// TIA Portal project "management parcare auto" (V17) (continued)
      ProcessValue <- "Status2"
   IOField "I/O field_77" at 1105,395 size 126x54; FormatPattern 9
      ProcessValue <- "Status3"
   IOField "I/O field_78" at 1105,445 size 126x54; FormatPattern 9
      ProcessValue <- "Status4"
   IOField "I/O field_79" at 1105,495 size 126x54; FormatPattern 9
      ProcessValue <- "Status5"
   IOField "I/O field_80" at 1105,545 size 126x54; FormatPattern 9
      ProcessValue <- "Status6"
   IOField "I/O field_81" at 1105,595 size 126x54; FormatPattern 9
      ProcessValue <- "Status7"
   IOField "I/O field_82" at 1105,645 size 126x54; FormatPattern 9
      ProcessValue <- "Status8"
   IOField "I/O field_83" at 1105,695 size 126x54; FormatPattern 9
      ProcessValue <- "Status9"
   IOField "I/O field_84" at 1105,745 size 126x54; FormatPattern 9
      ProcessValue <- "Status10"
   IOField "I/O field_85" at 1227,345 size 177x54; FormatPattern 9999999999999999999999999999999999999999
      ProcessValue <- "EntryTime2"
   IOField "I/O field_86" at 1227,395 size 177x54; FormatPattern 9999999999999999999999999999999999999999
      ProcessValue <- "EntryTime3"
   IOField "I/O field_87" at 1227,445 size 177x54; FormatPattern 9999999999999999999999999999999999999999
      ProcessValue <- "EntryTime4"
   IOField "I/O field_88" at 1227,495 size 177x54; FormatPattern 9999999999999999999999999999999999999999
      ProcessValue <- "EntryTime5"
   IOField "I/O field_89" at 1227,545 size 177x54; FormatPattern 9999999999999999999999999999999999999999
      ProcessValue <- "EntryTime6"
   IOField "I/O field_90" at 1227,595 size 177x54; FormatPattern 9999999999999999999999999999999999999999
      ProcessValue <- "EntryTime7"
   IOField "I/O field_91" at 1227,645 size 177x54; FormatPattern 9999999999999999999999999999999999999999
      ProcessValue <- "EntryTime8"
   IOField "I/O field_92" at 1227,695 size 177x54; FormatPattern 9999999999999999999999999999999999999999
      ProcessValue <- "EntryTime9"
   IOField "I/O field_93" at 1227,745 size 177x54; FormatPattern 9999999999999999999999999999999999999999
      ProcessValue <- "EntryTime10"
   IOField "I/O field_94" at 1400,344 size 165x54; FormatPattern 9999999999999999999999999999999999999999
      ProcessValue <- "EntryDate2"
   IOField "I/O field_95" at 1401,394 size 165x54; FormatPattern 9999999999999999999999999999999999999999
      ProcessValue <- "EntryDate3"
   IOField "I/O field_96" at 1401,444 size 165x54; FormatPattern 9999999999999999999999999999999999999999
      ProcessValue <- "EntryDate4"
   IOField "I/O field_97" at 1401,494 size 165x54; FormatPattern 9999999999999999999999999999999999999999
      ProcessValue <- "EntryDate5"
   IOField "I/O field_98" at 1401,545 size 165x54; FormatPattern 9999999999999999999999999999999999999999
      ProcessValue <- "EntryDate6"
   IOField "I/O field_99" at 1401,595 size 165x54; FormatPattern 9999999999999999999999999999999999999999
      ProcessValue <- "EntryDate7"
   IOField "I/O field_100" at 1401,645 size 165x54; FormatPattern 9999999999999999999999999999999999999999
      ProcessValue <- "EntryDate8"
   IOField "I/O field_101" at 1401,695 size 165x54; FormatPattern 9999999999999999999999999999999999999999
      ProcessValue <- "EntryDate9"
   IOField "I/O field_102" at 1401,745 size 165x54; FormatPattern 9999999999999999999999999999999999999999
      ProcessValue <- "EntryDate10"
   IOField "I/O field_103" at 1562,344 size 164x54; FormatPattern 9999999999999999999999999999999999999999
      ProcessValue <- "ExitTime2"
   IOField "I/O field_104" at 1562,394 size 164x54; FormatPattern 9999999999999999999999999999999999999999
      ProcessValue <- "ExitTime3"
   IOField "I/O field_105" at 1562,444 size 164x54; FormatPattern 9999999999999999999999999999999999999999
      ProcessValue <- "ExitTime4"
   IOField "I/O field_106" at 1562,494 size 164x54; FormatPattern 9999999999999999999999999999999999999999
      ProcessValue <- "ExitTime5"
   IOField "I/O field_107" at 1562,545 size 164x54; FormatPattern 9999999999999999999999999999999999999999
      ProcessValue <- "ExitTime6"
   IOField "I/O field_108" at 1562,595 size 164x54; FormatPattern 9999999999999999999999999999999999999999
      ProcessValue <- "ExitTime7"
   IOField "I/O field_109" at 1562,645 size 164x54; FormatPattern 9999999999999999999999999999999999999999
      ProcessValue <- "ExitTime8"
   IOField "I/O field_110" at 1562,695 size 164x54; FormatPattern 9999999999999999999999999999999999999999
      ProcessValue <- "ExitTime9"
   IOField "I/O field_111" at 1562,745 size 164x54; FormatPattern 9999999999999999999999999999999999999999
      ProcessValue <- "ExitTime10"
   IOField "I/O field_112" at 1723,344 size 163x54; FormatPattern 9999999999999999999999999999999999999999
      ProcessValue <- "ExitDate2"
   IOField "I/O field_113" at 1723,394 size 163x54; FormatPattern 9999999999999999999999999999999999999999
      ProcessValue <- "ExitDate3"
   IOField "I/O field_114" at 1723,444 size 163x54; FormatPattern 9999999999999999999999999999999999999999
      ProcessValue <- "ExitDate4"
   IOField "I/O field_115" at 1723,494 size 163x54; FormatPattern 9999999999999999999999999999999999999999
      ProcessValue <- "ExitDate5"
   IOField "I/O field_116" at 1723,544 size 163x54; FormatPattern 9999999999999999999999999999999999999999
      ProcessValue <- "ExitDate6"
   IOField "I/O field_117" at 1723,594 size 163x54; FormatPattern 9999999999999999999999999999999999999999
      ProcessValue <- "ExitDate7"
   IOField "I/O field_118" at 1723,644 size 163x54; FormatPattern 9999999999999999999999999999999999999999
      ProcessValue <- "ExitDate8"
   IOField "I/O field_119" at 1723,694 size 163x54; FormatPattern 9999999999999999999999999999999999999999
      ProcessValue <- "ExitDate9"
   IOField "I/O field_120" at 1723,744 size 163x54; FormatPattern 9999999999999999999999999999999999999999
      ProcessValue <- "ExitDate10"
   TextField "Text field_4" at 994,221 size 165x119; Text 'Car number'
   TextField "Text field_6" at 11,130 size 645x121; Text 'Temporar data'
   TextField "Text field_8" at 978,132 size 901x121; Text 'Permanent data'

screen "Statistics" 1920x1080
   on GenerateScreen: "Statistica_masini_total"()
   Button "Button_3" at 608,973 size 194x96; TextOff 'Statistics'
      on Press: ActivateScreen("Statistics", 0)
   Button "Button_8" at 408,973 size 194x96; TextOff 'Parking history'
      on Press: ActivateScreen("Parking history", 0)
   Button "Button_1" at 208,973 size 194x96; TextOff 'Alarms'
      on Press: ActivateScreen("Alarms", 0)
   Button "Button_2" at 9,972 size 194x96; TextOff 'Home / Ecran principal'
      on Press: ActivateScreen("Home", 0)
   GraphicView "Graphic view_2" at 28,12 size 394x64; Picture "Siemens_AG_logo.svg"
   Button "Button_4" at 1748,4 size 170x79; TextOff 'Exit / Iesire'
      on Press: StopRuntime(0)
   TextField "Text field_1" at 184,382 size 485x109; Text 'Number of cars:'
   TextField "Text field_2" at 794,230 size 49x81; Text 'Text'
   TextField "Text field_3" at 615,147 size 581x176; Text 'STATISTICS'
   TextField "Text field_4" at 164,210 size 1445x179; Text 'Choose a date(yy-mm-dd) to find out the number of cars on that day:'
   TextField "Text field_5" at 166,452 size 1589x179; Text 'Choose an interval to find out the number of cars in that period of time:'
   IOField "I/O field_1" at 316,328 size 178x62; FormatPattern ??????????
      on OnFinishInput: "Statistica_masini_zi"()
      ProcessValue <- "filtrare_dupa_data"
   IOField "I/O field_2" at 641,404 size 128x68; FormatPattern 99999
      ProcessValue <- "Numar_masini_ziuaX"
   TextField "Text field_6" at 512,561 size 26x62; Text '-'
   IOField "I/O field_4" at 312,569 size 188x62; FormatPattern ??????????
      ProcessValue <- "Interval1_date"
   IOField "I/O field_3" at 566,568 size 188x62; FormatPattern ??????????
      on OnFinishInput: "Statistica_masini_pe_interval"()
      ProcessValue <- "Interval2_date"
   TextField "Text field_7" at 166,621 size 485x109; Text 'Number of cars:'
   IOField "I/O field_5" at 615,647 size 128x68; FormatPattern 99999
      ProcessValue <- "nr_masini_interval"
   TextField "Text field_8" at 262,783 size 725x133; Text 'Total number of cars:'
   IOField "I/O field_6" at 1006,829 size 204x52; FormatPattern 9999999
      ProcessValue <- "nr_total_masini"

VB script "Insert_to_database"
   'RdyToLog= un tagg care se face 1 atunci cand butonul entry de pe HMI(nu runtime) este activat, devine trigger pentru a rula scriptul
   SmartTags("Verficare_rulareScriptInsr")=0
   If (SmartTags("RdyToLog")=True) And (SmartTags("04_DB_MarkersAuto_car status_1")=True Or SmartTags("04_DB_MarkersAuto_car status_2")=True Or SmartTags("04_DB_MarkersAuto_car status_3")=True Or SmartTags("04_DB_MarkersAuto_car status_4")=True Or SmartTags("04_DB_MarkersAuto_car status_5")=True Or SmartTags("04_DB_MarkersAuto_car status_6")=True Or SmartTags("04_DB_MarkersAuto_car status_7")=True Or SmartTags("04_DB_MarkersAuto_car status_8")=True Or SmartTags("04_DB_MarkersAuto_car status_9")=True Or SmartTags("04_DB_MarkersAuto_car status_10")=True ) Then
   
   Dim rs,con
   Dim nrMasina, statusMasina, oraIntrare,dataIntrare,oraIesire,dataIesire,dsValueEntry,dsValueExit
   
   
   'se ia nr de masina introdus de utilizator
   Set nrMasina= SmartTags("02_DB_HMI_Buttons_nr_masina")
   
   'se seteaza statusul masinii in functie de ce loc a ocupat
   If SmartTags("04_DB_MarkersAuto_car status_1")=True Then
   	statusMasina= 1
   End If
   
   If SmartTags("04_DB_MarkersAuto_car status_2")=True  Then
   	statusMasina=1
   End If
   
   If SmartTags("04_DB_MarkersAuto_car status_3")=True Then
   	statusMasina=1
   End If
   
   If SmartTags("04_DB_MarkersAuto_car status_4")=True Then
   	statusMasina=1
   End If
   
   If SmartTags("04_DB_MarkersAuto_car status_5")=True Then
   	statusMasina=1
   End If
   
   If SmartTags("04_DB_MarkersAuto_car status_6")=True Then
   	statusMasina=1
   End If
   
   If SmartTags("04_DB_MarkersAuto_car status_7")=True Then
   	statusMasina=1
   End If
   
   If SmartTags("04_DB_MarkersAuto_car status_8")=True Then
   	statusMasina=1
   End If
   
   If SmartTags("04_DB_MarkersAuto_car status_9")=True Then
   	statusMasina=1
   End If
   
   If  SmartTags("04_DB_MarkersAuto_car status_10")=True Then
   	statusMasina=1
   End If
   
   
   
   'Dim Timp
   'Timp = Time
   'Dim TimpStamp
   Dim dtsnow
   Dim dd, mm, yy, hh, nn, ss
   Dim DataValue, TimpValue
   
   'atunci cand se intra in parcare, se ia ora si data intrarii
   If SmartTags("11_DB_Inputs_i0.0")=True Then
   ' Obține data și ora curentă
   dtsnow = Now()
   dd = Right("00" & Day(dtsnow), 2)
   mm = Right("00" & Month(dtsnow), 2)
   yy = Year(dtsnow)
   
   hh = Right("00" & Hour(dtsnow), 2)
   nn = Right("00" & Minute(dtsnow), 2)
   ss = Right("00" & Second(dtsnow), 2)
   
   'Build the date string in the format yyyy-mm-dd
   dataIntrare = yy & "-" & mm & "-" & dd
   'Build the time string in the format hh:mm:ss
   oraIntrare = hh & ":" & nn & ":" & ss
   dsValueEntry=dataIntrare &" "& oraIntrare
   End If
   
   'atunci cand se plateste se ia ora si data iesirii
   If SmartTags("02_DB_HMI_Buttons_pay")=True Then
   ' Obține data și ora curentă
   dtsnow = Now()
   dd = Right("00" & Day(dtsnow), 2)
   mm = Right("00" & Month(dtsnow), 2)
   yy = Year(dtsnow)
   
   hh = Right("00" & Hour(dtsnow), 2)
   nn = Right("00" & Minute(dtsnow), 2)
   ss = Right("00" & Second(dtsnow), 2)
   
   'Build the date string in the format dd-mm-yyyy
   dataIesire = yy & "-" & mm & "-" & dd
   'Build the time string in the format hh:mm:ss
   oraIesire = hh & ":" & nn & ":" & ss
   dsValueExit=dataIesire & " " &oraIesire
   
   End If
   
   'conexiune baza de date si inserare
   Set con=CreateObject("adodb.connection")
   Set rs=CreateObject("adodb.recordset")
   
   con.open"Driver={MySQL ODBC 8.0 Unicode Driver};Server=localhost:3306;Database=parkingcar;User=root;Password=;Option=3;"
   Dim rezultate,rez
   rez="INSERT INTO parkingcar.permanent(NrInm,StatusMasina,OraIntrare,DataIntrare,OraIesire,DataIesire,DataOraEntry,DataOraExit) VALUES ('" & nrMasina & "', '" & statusMasina & "', '" & oraIntrare & "','" & dataIntrare & "','" & oraIesire & "','" & dataIesire & "', '" & dsValueEntry &"','"& dsValueExit &"')"
   rezultate= "INSERT INTO parkingcar.temporar(NrInm,StatusMasina,OraIntrare,DataIntrare,OraIesire,DataIesire,DataOraIntr,DataOraIesire) VALUES ('" & nrMasina & "', '" & statusMasina & "', '" & oraIntrare & "','" & dataIntrare & "','" & oraIesire & "','" & dataIesire & "', '" & dsValueEntry &"','"& dsValueExit &"')"
   rs.open rezultate,con
   rs.open rez,con
   con.Close
   End If
   
   SmartTags("Verficare_rulareScriptInsr")=1

VB script "EditDataRecord"
   'Tip:
   ' 1. Use the <CTRL+SPACE> or <CTRL+I> shortcut to open a list of all objects and functions
   ' 2. Write the code using the HMI Runtime object.
   '  Example: HmiRuntime.Screens("Screen_1").
   ' 3. Use the <CTRL+J> shortcut to create an object reference.
   'Write the code as of this position:
   
   
   If SmartTags("RdyToUpdate")=True Then
   Dim nrMasina,statusMasina, oraIesire,dataIesire
   Dim con,rs
   
   'se ia nr de masina folosit pentru a iesi din parcare
   Set nrMasina=SmartTags("02_DB_HMI_Buttons_nrMasina_iesire")
   
   If SmartTags("04_DB_MarkersAuto_car status_1")=False Then
   	statusMasina= 0
   End If
   
   If SmartTags("04_DB_MarkersAuto_car status_2")=False  Then
   	statusMasina=0
   End If
   
   If SmartTags("04_DB_MarkersAuto_car status_3")=False Then
   	statusMasina=0
   End If
   
   If SmartTags("04_DB_MarkersAuto_car status_4")=False Then
   	statusMasina=0
   End If
   
   If SmartTags("04_DB_MarkersAuto_car status_5")=False Then
   	statusMasina=0
   End If
   
   If SmartTags("04_DB_MarkersAuto_car status_6")=False Then
   	statusMasina=0
   End If
   
   If SmartTags("04_DB_MarkersAuto_car status_7")=False Then
   	statusMasina=0
   End If
   
   If SmartTags("04_DB_MarkersAuto_car status_8")=False Then
   	statusMasina=0
   End If
   
   If SmartTags("04_DB_MarkersAuto_car status_9")=False Then
   	statusMasina=0
   End If
   
   If  SmartTags("04_DB_MarkersAuto_car status_10")=False Then
   	statusMasina=0
   End If
   
   
   Dim dtsnow
   Dim dd, mm, yy, hh, nn, ss
   Dim DataValue, TimpValue,dsValueExit
   
   'atunci cand se plateste se ia ora si data iesirii
   If SmartTags("11_DB_Inputs_i1.0")=True Then
   ' Obține data și ora curentă
   dtsnow = Now()
   dd = Right("00" & Day(dtsnow), 2)
   mm = Right("00" & Month(dtsnow), 2)
   yy = Year(dtsnow)
   
   hh = Right("00" & Hour(dtsnow), 2)
   nn = Right("00" & Minute(dtsnow), 2)
   ss = Right("00" & Second(dtsnow), 2)
   
   'Build the date string in the format dd-mm-yyyy
   dataIesire = yy & "-" & mm & "-" & dd
   'Build the time string in the format hh:mm:ss
   oraIesire = hh & ":" & nn & ":" & ss
   dsValueExit=dataIesire &" " &oraIesire
   End If
   
   'conxiune baza de date si editare ora iesire si statusul
   Set con=CreateObject("adodb.connection")
   Set rs=CreateObject("adodb.recordset")
   
   con.open"Driver={MySQL ODBC 8.0 Unicode Driver};Server=localhost:3306;Database=parkingcar;User=root;Password=;Option=3;"
   Dim rezultate,rez
   rez="UPDATE parkingcar.permanent SET StatusMasina='" & statusMasina &"',OraIesire='" & oraIesire & "',DataIesire='" & dataIesire &"',DataOraExit='"& dsValueExit &"' WHERE NrInm='" & nrMasina &"' "
   rezultate= "UPDATE parkingcar.temporar SET StatusMasina='" & statusMasina &"',OraIesire='" & oraIesire & "',DataIesire='" & dataIesire &"', DataOraIesire='"& dsValueExit &"' WHERE NrInm='" & nrMasina &"' "
   rs.open rezultate,con
   rs.open rez,con
   con.Close
   
   End If

VB script "Delete_from_database"
   'Tip:
   ' 1. Use the <CTRL+SPACE> or <CTRL+I> shortcut to open a list of all objects and functions
   ' 2. Write the code using the HMI Runtime object.
   '  Example: HmiRuntime.Screens("Screen_1").
   ' 3. Use the <CTRL+J> shortcut to create an object reference.
   'Write the code as of this position:
   
   If SmartTags("RdyToDelete")=True Then
   	
   Dim con,rs
   
   Set con=CreateObject("adodb.connection")
   Set rs=CreateObject("adodb.recordset")
   
   con.open"Driver={MySQL ODBC 8.0 Unicode Driver};Server=localhost:3306;Database=parkingcar;User=root;Password=;Option=3;"
   Dim rezultate
   rezultate= "DELETE FROM parkingcar.temporar WHERE StatusMasina= '0'"
   rs.open rezultate,con
   con.Close
   End If

VB script "Statistica_masini_zi"
   'Tip:
   ' 1. Use the <CTRL+SPACE> or <CTRL+I> shortcut to open a list of all objects and functions
   ' 2. Write the code using the HMI Runtime object.
   '  Example: HmiRuntime.Screens("Screen_1").
   ' 3. Use the <CTRL+J> shortcut to create an object reference.
   'Write the code as of this position:
   
   Dim con,rs 
   Set con=CreateObject("ADODB.Connection")
   Set rs= CreateObject("adodb.recordset")
   
   con.Open "DRIVER={MySQL ODBC 8.0 Unicode Driver};Server=localhost:3306;Database=parkingcar;User=root;Password=;Option=3;"
   rs.open "SELECT  COUNT(* ) AS NumarMasini FROM permanent WHERE DataIntrare = '" & SmartTags("filtrare_dupa_data")&"' ",con
   SmartTags("Numar_masini_ziuaX")=rs.Fields(0)
   Set con=Nothing

VB script "Statistica_masini_pe_interval"
   'Tip:
   ' 1. Use the <CTRL+SPACE> or <CTRL+I> shortcut to open a list of all objects and functions
   ' 2. Write the code using the HMI Runtime object.
   '  Example: HmiRuntime.Screens("Screen_1").
   ' 3. Use the <CTRL+J> shortcut to create an object reference.
   'Write the code as of this position:
   Dim con,rs 
   Set con=CreateObject("ADODB.Connection")
   Set rs= CreateObject("adodb.recordset")
   
   con.Open "DRIVER={MySQL ODBC 8.0 Unicode Driver};Server=localhost:3306;Database=parkingcar;User=root;Password=;Option=3;"
   rs.open "SELECT  COUNT(* ) AS NumarMasini FROM permanent WHERE DataIntrare >= '" & SmartTags("Interval1_date") &"' AND DataIntrare <= '" & SmartTags("Interval2_date") &"' ",con
   SmartTags("nr_masini_interval")=rs.Fields(0)

VB script "Statistica_masini_total"
   'Tip:
   ' 1. Use the <CTRL+SPACE> or <CTRL+I> shortcut to open a list of all objects and functions
   ' 2. Write the code using the HMI Runtime object.
   '  Example: HmiRuntime.Screens("Screen_1").
   ' 3. Use the <CTRL+J> shortcut to create an object reference.
   'Write the code as of this position:
   
   Dim con,rs 
   Set con=CreateObject("ADODB.Connection")
   Set rs= CreateObject("adodb.recordset")
   
   con.Open "DRIVER={MySQL ODBC 8.0 Unicode Driver};Server=localhost:3306;Database=parkingcar;User=root;Password=;Option=3;"
   rs.open "SELECT  COUNT(* ) AS NumarMasini FROM permanent",con
   SmartTags("nr_total_masini")=rs.Fields(0)

VB script "Read_fromTEMP"
   'Tip:
   ' 1. Use the <CTRL+SPACE> or <CTRL+I> shortcut to open a list of all objects and functions
   ' 2. Write the code using the HMI Runtime object.
   '  Example: HmiRuntime.Screens("Screen_1").
   ' 3. Use the <CTRL+J> shortcut to create an object reference.
   'Write the code as of this position:
   Dim con,rs
   ' Creează obiectul pentru conexiunea la bază de date
   Set con = CreateObject("ADODB.Connection")
   Set rs=CreateObject("adodb.recordset")
    
   ' Deschide conexiunea la bază de date
   con.Open "DRIVER={MySQL ODBC 8.0 Unicode Driver};Server=localhost:3306;Database=parkingcar;User=root;Password=;Option=3;"
   rs.open "SELECT * FROM temporar ORDER BY NrInm ASC ",con
   rs.MoveFirst
   Dim i
   i=1
   While Not rs.EOF
   SmartTags("NrMasina"& i)=rs.Fields("NrInm")
   SmartTags("CarStatus"& i)=rs.Fields("StatusMasina")
   SmartTags("OraIntrare"& i)=rs.Fields("DataOraIntr")
   SmartTags("DataIntrare"& i)=rs.Fields("DataOraIntr")
   rs.MoveNext
   i=i+1
   Wend
   
   If rs.EOF Then
   	rs.Close
   	con.Close
   End If

VB script "Read_fromPerm"
   'Tip:
   ' 1. Use the <CTRL+SPACE> or <CTRL+I> shortcut to open a list of all objects and functions
   ' 2. Write the code using the HMI Runtime object.
   '  Example: HmiRuntime.Screens("Screen_1").
   ' 3. Use the <CTRL+J> shortcut to create an object reference.
   'Write the code as of this position:
   
   Dim con,rs
   ' Creează obiectul pentru conexiunea la bază de date
   Set con = CreateObject("ADODB.Connection")
   Set rs=CreateObject("adodb.recordset")
    Dim exittime
    exittime="00-00-00 00:00:00"
   ' Deschide conexiunea la bază de date
   con.Open "DRIVER={MySQL ODBC 8.0 Unicode Driver};Server=localhost:3306;Database=parkingcar;User=root;Password=;Option=3;"
   rs.open "SELECT * FROM permanent ORDER BY DataIntrare DESC",con
   rs.MoveFirst
   Dim i
   'Please replace all sequences which are enclosed with '_' by your own code.
   For  i= 1 To 10
   SmartTags("CarNumber"& i)=rs.Fields("NrInm")
   SmartTags("Status"& i)=rs.Fields("StatusMasina")
   SmartTags("EntryTime"& i)=rs.Fields("DataOraEntry")
   SmartTags("EntryDate"& i)=rs.Fields("DataOraEntry")
   Dim value
   value=rs.Fields("DataOraExit")
   If IsNull(value) Then
   	SmartTags("ExitTime" & i)=0
   	SmartTags("ExitDate" & i)=0
   Else
   	SmartTags("ExitTime" & i)=CDate(rs.Fields("DataOraExit"))
   	SmartTags("ExitDate" & i)=CDate(rs.Fields("DataOraExit"))
   End If
   rs.MoveNext
   Next
   
   rs.Close
   con.Close
*)

(* ===== HMI "HMI_RT_2" =====
system functions are stored by id; their names below are inferred from use
connection "HMI_Connection_1": ETHERNET, SMART_S7_1500_OMS

HMI tags "Default tag table"
   "02_DB_HMI_Buttons_pay" : Bool = PLC "02_DB_HMI_Buttons".pay, 1 s
   "04_DB_MarkersAuto_remaining parking lots" : Int = PLC "04_DB_MarkersAuto"."remaining parking lots", 1 s
   "02_DB_HMI_Buttons_nr_masina" : String[254] = PLC "02_DB_HMI_Buttons".nrMasina_intrare, 1 s
   "02_DB_HMI_Buttons_nrMasina_iesire" : String[254] = PLC "02_DB_HMI_Buttons".nrMasina_iesire, 1 s
   "11_DB_Inputs_i0.1" : Bool = PLC "11_DB_Inputs"."i0.1", 1 s
   "11_DB_Inputs_i0.2" : Bool = PLC "11_DB_Inputs"."i0.2", 1 s
   "11_DB_Inputs_i0.3" : Bool = PLC "11_DB_Inputs"."i0.3", 1 s
   "11_DB_Inputs_i0.4" : Bool = PLC "11_DB_Inputs"."i0.4", 1 s
   "11_DB_Inputs_i0.5" : Bool = PLC "11_DB_Inputs"."i0.5", 1 s
   "11_DB_Inputs_i0.6" : Bool = PLC "11_DB_Inputs"."i0.6", 1 s
   "11_DB_Inputs_i0.7" : Bool = PLC "11_DB_Inputs"."i0.7", 1 s
   "11_DB_Inputs_i1.1" : Bool = PLC "11_DB_Inputs"."i1.1", 1 s
   "11_DB_Inputs_i1.2" : Bool = PLC "11_DB_Inputs"."i1.2", 1 s
   "11_DB_Inputs_i1.3" : Bool = PLC "11_DB_Inputs"."i1.3", 1 s
   "02_DB_HMI_Buttons_Parking lot 1" : Bool = PLC "02_DB_HMI_Buttons"."Parking lot 1", 1 s
   "02_DB_HMI_Buttons_Parking lot 2" : Bool = PLC "02_DB_HMI_Buttons"."Parking lot 2", 1 s
   "02_DB_HMI_Buttons_Parking lot 3" : Bool = PLC "02_DB_HMI_Buttons"."Parking lot 3", 1 s
   "02_DB_HMI_Buttons_Parking lot 4" : Bool = PLC "02_DB_HMI_Buttons"."Parking lot 4", 1 s
   "02_DB_HMI_Buttons_Parking lot 5" : Bool = PLC "02_DB_HMI_Buttons"."Parking lot 5", 1 s
   "02_DB_HMI_Buttons_Parking lot 6" : Bool = PLC "02_DB_HMI_Buttons"."Parking lot 6", 1 s
   "02_DB_HMI_Buttons_Parking lot 7" : Bool = PLC "02_DB_HMI_Buttons"."Parking lot 7", 1 s
   "02_DB_HMI_Buttons_Parking lot 8" : Bool = PLC "02_DB_HMI_Buttons"."Parking lot 8", 1 s
   "02_DB_HMI_Buttons_Parking lot 9" : Bool = PLC "02_DB_HMI_Buttons"."Parking lot 9", 1 s
   "02_DB_HMI_Buttons_Parking lot 10" : Bool = PLC "02_DB_HMI_Buttons"."Parking lot 10", 1 s
   "11_DB_Inputs_i0.0" : Bool = PLC "11_DB_Inputs"."i0.0", 1 s
   "11_DB_Inputs_i1.0" : Bool = PLC "11_DB_Inputs"."i1.0", 1 s

HMI tags "Alarms"
   "Alarma_full" : Word = PLC "08_DB_Alarms".Full AT %DB1.DBW0, 1 s
   "Alarma_loc neselectat" : Word = PLC "08_DB_Alarms".Parking_lot_empty AT %DB1.DBW0, 1 s
   "Alarma_barieraIntr_nu" : Word = PLC "08_DB_Alarms".EntryBarrierNotWorking AT %DB1.DBW0, 1 s
   "Alarma_barieraIesire_nu" : Word = PLC "08_DB_Alarms".ExitBarrierNotWorking AT %DB1.DBW0, 1 s

discrete alarms
   1: 'The car park is at maximum capacity. You have nowhere to park! / Parcarea este la capacitatea maxima. Nu aveti unde sa parcati!', class Warnings, trigger "Alarma_full" bit 0
   2: 'No parking space has been selected. Please select a free parking spot! / Niciun loc de parcare nu a fost selectat. Te rugam sa selectezi un loc liber!', class Warnings, trigger "Alarma_loc neselectat" bit 0
   3: 'The entry barrier does not work! Call the operator! / Bariera de la intrare nu functioneaza! Chemati un operator!', class Errors, trigger "Alarma_barieraIntr_nu" bit 0
   4: 'The exit barrier does not work! Call the operator! / Bariera de la iesire nu functuioneaza! Chemati un operator!', class Errors, trigger "Alarma_barieraIesire_nu" bit 0

screen "Exit" 800x480
   TextField "Text field_1" at 190,86 size 408x91; Text 'Car park / Parcare auto'
   Button "Button_1" at 279,294 size 213x80; TextOff 'Pay / Plateste'
      on Press: SetBit("02_DB_HMI_Buttons_pay")
      on Release: ResetBit("02_DB_HMI_Buttons_pay"); ActivateScreen("root screen", 0)
   GraphicView "Graphic view_1" at 9,9 size 198x51; Picture "Siemens_AG_logo.svg"
   Button "Button_2" at 646,414 size 141x60; TextOff 'Exit / Iesire'; Authorization "operator"
      on Press: StopRuntime(0); function_a2a04561()
   GraphicView "Graphic view_2" at 648,430 size 36x30; Picture "Graphic_1"
   DateTimeField "Date/time field_1" at 568,16 size 219x32
   Button "Button_3" at 161,415 size 141x60; TextOff 'Alarms / Alarme'
      on Press: ActivateScreen("Alarms", 0)
   IOField "I/O field_1" at 651,127 size 124x44; FormatPattern s99999
      ProcessValue <- "04_DB_MarkersAuto_remaining parking lots"
   TextField "Text field_13" at 59,204 size 366x50; Text 'Enter the registration number of the car and then you can pay: Introduceti numarul de inmatriculare si dupa puteti sa platiti!'
   IOField "I/O field_3" at 381,230 size 165x38; FormatPattern ????????
      ProcessValue <- "02_DB_HMI_Buttons_nrMasina_iesire"
   Button "Button_4" at 9,415 size 141x60; TextOff 'Back / Inapoi'
      on Press: ActivateScreen("root screen", 0)
   Ellipse "Ellipse_1" at 748,248 size 39x32
      Appearance <- "11_DB_Inputs_i0.0"
   Ellipse "Ellipse_2" at 750,324 size 39x32
      Appearance <- "11_DB_Inputs_i1.0"
   TextField "Text field_3" at 662,214 size 122x23; Text 'Entry sensor / Senzor intrare'
   TextField "Text field_4" at 668,296 size 111x23; Text 'Exit sensor / Senzor iesire'
   Button "Button_5" at 633,247 size 109x32; TextOff 'ON/OFF / Pornit/Oprit'
      on Press: InvertBit("11_DB_Inputs_i0.0")
   Button "Button_6" at 636,325 size 106x32; TextOff 'ON/OFF / Pornit/Oprit'
      on Press: InvertBit("11_DB_Inputs_i1.0")
   TextField "Text field_2" at 716,93 size 65x29; Text 'Free: / Liber:'

screen "Alarms" 800x480
   TextField "Text field_1" at 271,67 size 226x91; Text 'Alarms / Alarme'
   GraphicView "Graphic view_1" at 9,9 size 198x51; Picture "Siemens_AG_logo.svg"
   Button "Button_2" at 646,414 size 141x60; TextOff 'Exit / Iesire'; Authorization "operator"
      on Press: StopRuntime(0); function_a2a04561()
   GraphicView "Graphic view_2" at 642,430 size 36x30; Picture "Graphic_1"
   DateTimeField "Date/time field_1" at 568,16 size 219x32
   Button "Button_3" at 9,415 size 141x60; TextOff 'Back / Inapoi'
      on Press: ActivateScreen("root screen", 0)
   AlarmView "Alarm view_1" at 40,155 size 725x253

screen "Entry" 800x480
   TextField "Text field_13" at 4,71 size 308x94; Text 'Enter the registration number of the car and then select a free space: Introduceti nr. de inmatriculare si dupa selectati un loc liber:'
   Rectangle "Rectangle_10" at 450,279 size 115x101
      Appearance <- "11_DB_Inputs_i1.2"
   Rectangle "Rectangle_9" at 569,279 size 115x101
      Appearance <- "11_DB_Inputs_i1.3"
   Rectangle "Rectangle_8" at 331,279 size 115x101
      Appearance <- "11_DB_Inputs_i1.1"
   Rectangle "Rectangle_7" at 211,280 size 115x99
      Appearance <- "11_DB_Inputs_i0.7"
   Rectangle "Rectangle_6" at 92,279 size 115x101
      Appearance <- "11_DB_Inputs_i0.6"
   Rectangle "Rectangle_5" at 569,172 size 115x103
      Appearance <- "11_DB_Inputs_i0.5"
   Rectangle "Rectangle_4" at 450,172 size 115x103
      Appearance <- "11_DB_Inputs_i0.4"
   Rectangle "Rectangle_3" at 330,172 size 115x103
      Appearance <- "11_DB_Inputs_i0.3"
   Rectangle "Rectangle_2" at 211,172 size 115x103
      Appearance <- "11_DB_Inputs_i0.2"
   Rectangle "Rectangle_1" at 92,172 size 115x103
      Appearance <- "11_DB_Inputs_i0.1"
   TextField "Text field_1" at 372,98 size 238x47; Text 'Car park / Parcare auto'
   GraphicView "Graphic view_1" at 9,9 size 198x51; Picture "Siemens_AG_logo.svg"
   Button "Button_2" at 646,414 size 141x60; TextOff 'Exit / Iesire'; Authorization "operator"
      on Press: StopRuntime(0); function_a2a04561()
   GraphicView "Graphic view_2" at 643,430 size 36x30; Picture "Graphic_1"
   DateTimeField "Date/time field_1" at 568,16 size 219x32
   Button "Button_3" at 160,416 size 141x60; TextOff 'Alarms / Alarme'
      on Press: ActivateScreen("Alarms", 0)
   IOField "I/O field_1" at 689,103 size 92x44; FormatPattern s99999
      ProcessValue <- "04_DB_MarkersAuto_remaining parking lots"
   Group "Group" at 90,169 size 596x213
   TextField "Text field_3" at 122,231 size 51x47; Text '01'
   TextField "Text field_4" at 242,231 size 51x47; Text '02'
   TextField "Text field_5" at 361,231 size 51x47; Text '03'
   TextField "Text field_6" at 482,231 size 51x47; Text '04'
   TextField "Text field_7" at 602,231 size 51x47; Text '05'
   TextField "Text field_8" at 122,335 size 51x47; Text '06'
   TextField "Text field_9" at 242,335 size 51x47; Text '07'
   TextField "Text field_10" at 361,335 size 51x47; Text '08'
   TextField "Text field_11" at 482,335 size 51x47; Text '09'
   TextField "Text field_12" at 602,335 size 51x47; Text '10'
   Button "Button_1" at 101,177 size 100x41; TextOff 'Parking lot no.1 Loc parcare nr.1'
      on Press: SetBit("02_DB_HMI_Buttons_Parking lot 1")
      on Release: ResetBit("02_DB_HMI_Buttons_Parking lot 1"); ActivateScreen("root screen", 0)
      Visibility <- "11_DB_Inputs_i0.1"
      Appearance <- "02_DB_HMI_Buttons_Parking lot 1"
   Button "Button_4" at 217,177 size 100x41; TextOff 'Parking lot no.2 Loc parcare nr.2'
      on Press: SetBit("02_DB_HMI_Buttons_Parking lot 2")
      on Release: ResetBit("02_DB_HMI_Buttons_Parking lot 2"); ActivateScreen("root screen", 0)
      Visibility <- "11_DB_Inputs_i0.2"
      Appearance <- "02_DB_HMI_Buttons_Parking lot 2"
   Button "Button_5" at 339,177 size 100x41; TextOff 'Parking lot no.3 Loc parcare nr.3'
      on Press: SetBit("02_DB_HMI_Buttons_Parking lot 3")
      on Release: ResetBit("02_DB_HMI_Buttons_Parking lot 3"); ActivateScreen("root screen", 0)
      Visibility <- "11_DB_Inputs_i0.3"
      Appearance <- "02_DB_HMI_Buttons_Parking lot 3"
   Button "Button_6" at 459,177 size 100x41; TextOff 'Parking lot no.4 Loc parcare nr.4'
      on Press: SetBit("02_DB_HMI_Buttons_Parking lot 4")
      on Release: ResetBit("02_DB_HMI_Buttons_Parking lot 4"); ActivateScreen("root screen", 0)
      Visibility <- "11_DB_Inputs_i0.4"
      Appearance <- "02_DB_HMI_Buttons_Parking lot 4"
   Button "Button_7" at 579,177 size 100x41; TextOff 'Parking lot no.5 Loc parcare nr.5'
      on Press: SetBit("02_DB_HMI_Buttons_Parking lot 5")
      on Release: ResetBit("02_DB_HMI_Buttons_Parking lot 5"); ActivateScreen("root screen", 0)
      Visibility <- "11_DB_Inputs_i0.5"
      Appearance <- "02_DB_HMI_Buttons_Parking lot 5"
   Button "Button_8" at 101,285 size 100x41; TextOff 'Parking lot no.6 Loc parcare nr.6'
      on Press: SetBit("02_DB_HMI_Buttons_Parking lot 6")
      on Release: ResetBit("02_DB_HMI_Buttons_Parking lot 6"); ActivateScreen("root screen", 0)
      Visibility <- "11_DB_Inputs_i0.6"
      Appearance <- "02_DB_HMI_Buttons_Parking lot 6"
   Button "Button_9" at 219,285 size 100x41; TextOff 'Parking lot no.7 Loc parcare nr.7'
      on Press: SetBit("02_DB_HMI_Buttons_Parking lot 7")
      on Release: ResetBit("02_DB_HMI_Buttons_Parking lot 7"); ActivateScreen("root screen", 0)
      Visibility <- "11_DB_Inputs_i0.7"
      Appearance <- "02_DB_HMI_Buttons_Parking lot 7"
   Button "Button_10" at 339,285 size 100x41; TextOff 'Parking lot no.8 Loc parcare nr.8'
      on Press: SetBit("02_DB_HMI_Buttons_Parking lot 8")
      on Release: ResetBit("02_DB_HMI_Buttons_Parking lot 8"); ActivateScreen("root screen", 0)
      Visibility <- "11_DB_Inputs_i1.1"
      Appearance <- "02_DB_HMI_Buttons_Parking lot 8"
   Button "Button_11" at 459,285 size 100x41; TextOff 'Parking lot no.9 Loc parcare nr.9'
      on Press: SetBit("02_DB_HMI_Buttons_Parking lot 9")
      on Release: ResetBit("02_DB_HMI_Buttons_Parking lot 9"); ActivateScreen("root screen", 0)
      Visibility <- "11_DB_Inputs_i1.2"
      Appearance <- "02_DB_HMI_Buttons_Parking lot 9"
   Button "Button_12" at 579,285 size 100x41; TextOff 'Parking lot no.10 Loc parcare nr.10'
      on Press: SetBit("02_DB_HMI_Buttons_Parking lot 10")
      on Release: ResetBit("02_DB_HMI_Buttons_Parking lot 10"); ActivateScreen("root screen", 0)
      Visibility <- "11_DB_Inputs_i1.3"
      Appearance <- "02_DB_HMI_Buttons_Parking lot 10"
   Button "Button_13" at 9,415 size 141x60; TextOff 'Back / Inapoi'
      on Press: ActivateScreen("root screen", 0)
   IOField "I/O field_2" at 160,126 size 98x42; FormatPattern ????????
      ProcessValue <- "02_DB_HMI_Buttons_nr_masina"
   Ellipse "Ellipse_1" at 717,200 size 39x32
      Appearance <- "11_DB_Inputs_i0.0"
   Ellipse "Ellipse_2" at 719,325 size 39x32
      Appearance <- "11_DB_Inputs_i1.0"
   TextField "Text field_14" at 683,161 size 106x42; Text 'Entry sensor Senzor intrare'
   TextField "Text field_15" at 693,288 size 95x42; Text 'Exit sensor Senzor iesire'
   Button "Button_14" at 691,237 size 105x32; TextOff 'ON/OFF / Pornit/Oprit'
      on Press: InvertBit("11_DB_Inputs_i0.0")
   Button "Button_15" at 689,361 size 103x32; TextOff 'ON/OFF / Pornit/Oprit'
      on Press: InvertBit("11_DB_Inputs_i1.0")
   TextField "Text field_2" at 717,75 size 65x29; Text 'Free: / Liber:'

screen "root screen" 800x480
   TextField "Text field_1" at 236,78 size 408x91; Text 'Car park / Parcare auto'
   Button "Button_1" at 299,192 size 213x80; TextOff 'Entry / Intrare'
      on Press: ActivateScreen("Entry", 0)
      Visibility <- "Alarma_full"
   GraphicView "Graphic view_1" at 9,9 size 198x51; Picture "Siemens_AG_logo.svg"
   Button "Button_2" at 644,414 size 143x60; TextOff 'Exit / Iesire'; Authorization "operator"
      on Press: StopRuntime(0)
   GraphicView "Graphic view_2" at 641,430 size 36x30; Picture "Graphic_1"
   DateTimeField "Date/time field_1" at 568,16 size 219x32
   Button "Button_3" at 9,415 size 141x60; TextOff 'Alarms / Alarme'
      on Press: ActivateScreen("Alarms", 0)
   IOField "I/O field_1" at 651,104 size 124x44; FormatPattern s99999
      ProcessValue <- "04_DB_MarkersAuto_remaining parking lots"
   Button "Button_4" at 298,293 size 213x80; TextOff 'Exit / Iesire'
      on Press: ActivateScreen("Exit", 0)
   Ellipse "Ellipse_1" at 748,206 size 39x32
      Appearance <- "11_DB_Inputs_i0.0"
   Ellipse "Ellipse_2" at 750,282 size 39x32
      Appearance <- "11_DB_Inputs_i1.0"
   TextField "Text field_3" at 662,177 size 122x23; Text 'Entry sensor / Senzor intrare'
   TextField "Text field_4" at 668,254 size 111x23; Text 'Exit sensor / Senzor iesire'
   Button "Button_5" at 632,207 size 110x30; TextOff 'ON/OFF / Pornit/Oprit'
      on Press: InvertBit("11_DB_Inputs_i0.0")
   Button "Button_6" at 631,283 size 111x32; TextOff 'ON/OFF / Pornit/Oprit'
      on Press: InvertBit("11_DB_Inputs_i1.0")
   Rectangle "Rectangle_1" at 188,168 size 419x104
      Visibility <- "Alarma_full"
   TextField "Text field_5" at 203,199 size 404x54; Text 'Maximum capacity has been reached! No more parking lots available! Capacitatea maxima a fost atinsa. Nu mai sunt locuri de parcare libere!'
      Visibility <- "Alarma_full"
   GraphicView "Graphic view_3" at 187,179 size 36x30; Picture "Graphic_6"
      Visibility <- "Alarma_full"
   Button "Button_7" at 9,70 size 67x38; TextOff 'Text'; PictureOff "english_1"
      on Click: function_fb9197e8(L en-US)
   Button "Button_8" at 91,70 size 67x38; TextOff 'Text'; PictureOff "download (2)"
      on Click: function_fb9197e8(L ro-RO)
   TextField "Text field_2" at 717,75 size 65x29; Text 'Free: / Liber:'
*)